        [10]   // MV 36,TEMPERATURE SETPOINT E. 1/10 DEGREE 'C'
        [12]   // MV 36,TEMPERATURE SETPOINT F. 1/10 DEGREE 'C'
        [14]   // MV 36,TEMPERATURE SETPOINT G. 1/10 DEGREE 'C'
        [13]   // MV 36,TEMPERATURE BREAKPOINT G. TIME 1/10 HOURS(ALWAYS=0)
        [15].2   // MV 36,PLC TO FOLLOW RAMP Breakpoints A to B
        [30].6   // MV 36,Current vessel cold cond.temp.reached
        [27]   // MV 36,CURRENT ELAPSED HOURS *10
        [30].5   // MV 36,Current vessel deferred chilling temp.high flag
        [1]   // MV 36,TEMPERATURE BREAKPOINT A. TIME 1/10 HOURS(ALWAYS=0)
        [29].1   // MV 36,Current vessel deferred chilling enabled flag
        [30].0   // MV 36,Cooling Valve to open
        [3]   // MV 36,TEMPERATURE BREAKPOINT B. TIME 1/10 HOURS(ALWAYS=0)
        [5]   // MV 36,TEMPERATURE BREAKPOINT C. TIME 1/10 HOURS(ALWAYS=0)
        [7]   // MV 36,TEMPERATURE BREAKPOINT D. TIME 1/10 HOURS(ALWAYS=0)
        [9]   // MV 36,TEMPERATURE BREAKPOINT E. TIME 1/10 HOURS(ALWAYS=0)
        [22]   // MV 36,Current FV total residence time
        [15].7   // MV 36,PC>PLC Rousing enabled
        [29].0   // MV 36,PC TO SAVE TEMPERATURE DATA
        [43]   // MV 36,Current vessel powder type
        [44]   // MV 36,Current vessel powder amount
        [15].3   // MV 36,PLC TO USE CONE COOLING JACKET
        [25]   // MV 36,ACTUAL TEMPERATURE -DEGREES 'C'*10
        [15]   // MV 36,FLAGS-PROFILE CONTROL
        [26]   // MV 36,Calculated Setpoint 1/10 degrees C
        [20]   // MV 36,Current FV warm conditioning time
        [29]   // MV 36,FLAGS - PLC CONTROL
        [30].1   // MV 36,Rouser required
        [28]   // MV 36,CURRENT VOLUME HL*10
   MV_N151 : INT[50] := ([0] := 347, [2] := 100, [3] := 1200, [4] := 100, [5] := 1680, [6] := -15, [7] := 5280, [8] := -15, [9] := 7210, [10] := -15, [11] := 8340, [12] := -15, [13] := 32767, [14] := -15, [15] := 164, [17] := -32767, [18] := -32767, [19] := 1680, [20] := 1200, [21] := 2981, [22] := 6282, [23] := 1, [24] := 13, [25] := -12, [26] := -15, [27] := 4630, [30] := 123, [32] := 2, [34] := 2, [40] := 2);   // MV 47, CURRENT FV DATA
        [24]   // MV 47,Phase 0=off 8=Wait yeast 9=Wait Fill 10=Maturation 11to16=Conditioning
        [15].9   // MV 47,Current vessel deferred chilling manual override
        [15].4   // MV 47,Profile Control Flags : This is a Maturation Profile
        [30].3   // MV 47,Current vessel deferred chilling active
        [15].5   // MV 47,Profile Control Flags : This is a Conditioning Profile
        [11]   // MV 47,TEMPERATURE BREAKPOINT F. TIME 1/10 HOURS(ALWAYS=0)
        [13]   // MV 47,TEMPERATURE BREAKPOINT G. TIME 1/10 HOURS(ALWAYS=0)
        [16].1   // MV 47,Profile control flag Hold at B.P B
        [16].2   // MV 47,Profile control flag Hold at B.P C
        [16].3   // MV 47,Profile control flag Hold at B.P D
        [30].5   // MV 47,Current vessel deferred chilling temp.high flag
        [36]   // MV 47,Current vessel time to deferred chlling start (hrs.x10)
        [16].4   // MV 47,Profile control flag Hold at B.P E
        [16].5   // MV 47,Profile control flag Hold at B.P F
        [16].6   // MV 47,Profile control flag Hold at B.P G
        [0]   // MV 47,FV SYSTEM WORKING BUFFER VESSEL NUMBER
        [21]   // MV 47,Current vessel cold conditioning time
        [2]   // MV 47,TEMPERATURE SETPOINT A. 1/10 DEGREE 'C'
        [30].4   // MV 47,Current vessel final temp.reached
        [4]   // MV 47,TEMPERATURE SETPOINT B. 1/10 DEGREE 'C'
        [6]   // MV 47,TEMPERATURE SETPOINT C. 1/10 DEGREE 'C'
        [8]   // MV 47,TEMPERATURE SETPOINT D. 1/10 DEGREE 'C'
        [40]   // MV 47,Vessel RoutingStatus 0=Clean,1=Filling,2= Beer,3=Packng1,4=Pac kng2,5=Packng3,6=Ven ting,7=Dirty,8=CIP
        [10]   // MV 47,TEMPERATURE SETPOINT E. 1/10 DEGREE 'C'
        [1]   // MV 47,TEMPERATURE BREAKPOINT A. TIME 1/10 HOURS(ALWAYS=0)
        [12]   // MV 47,TEMPERATURE SETPOINT F. 1/10 DEGREE 'C'
        [14]   // MV 47,TEMPERATURE SETPOINT G. 1/10 DEGREE 'C'
        [29].1   // MV 47,Current vessel deferred chilling enabled flag
        [15].2   // MV 47,PLC TO FOLLOW RAMP Breakpoints A to B
        [30].6   // MV 47,Current vessel cold cond.temp.reached
        [3]   // MV 47,TEMPERATURE BREAKPOINT B. TIME 1/10 HOURS(ALWAYS=0)
        [5]   // MV 47,TEMPERATURE BREAKPOINT C. TIME 1/10 HOURS(ALWAYS=0)
        [27]   // MV 47,CURRENT ELAPSED HOURS *10
        [30].0   // MV 47,Cooling Valve to open
        [7]   // MV 47,TEMPERATURE BREAKPOINT D. TIME 1/10 HOURS(ALWAYS=0)
        [9]   // MV 47,TEMPERATURE BREAKPOINT E. TIME 1/10 HOURS(ALWAYS=0)
        [22]   // MV 47,Current FV total residence time
        [15].7   // MV 47,PC>PLC Rousing enabled
        [43]   // MV 47,Current vessel powder type
        [29].0   // MV 47,PC TO SAVE TEMPERATURE DATA
        [15].3   // MV 47,PLC TO USE CONE COOLING JACKET
        [44]   // MV 47,Current vessel powder amount
        [25]   // MV 47,ACTUAL TEMPERATURE -DEGREES 'C'*10
        [15]   // MV 47,FLAGS-PROFILE CONTROL
        [26]   // MV 47,Calculated Setpoint 1/10 degrees C
        [20]   // MV 47,Current FV warm conditioning time
        [29]   // MV 47,FLAGS - PLC CONTROL
        [30].1   // MV 47,Rouser required
        [28]   // MV 47,CURRENT VOLUME HL*10
   MV_N15_63_0_OutputBit : BOOL;
   MV_N190 : INT[255] := ([0] := 1, [2] := 2, [3] := 2, [4] := 7, [5] := 2, [6] := 2, [7] := 2, [8] := 2, [9] := 2, [10] := 7, [11] := 7, [12] := 7, [13] := 2, [100] := 1, [101] := 2048, [102] := 10, [103] := 14, [105] := 13, [106] := 10, [107] := 15, [108] := 10, [109] := 10, [113] := 10, [200] := 8194, [201] := -16384, [203] := 20, [204] := 11, [205] := 137, [206] := 100, [209] := 23, [215] := 14641, [216] := 11826, [217] := 13873, [218] := 11832, [219] := 12338, [220] := 13102, [221] := 52);   // Original N File From SLC, No Description Available
        [200].0   // Heartbeat Fault
        [101].0   // MV36 Rouser On to Remote I/O on MV Routing PLC
        [101].1   // MV37 Rouser On to Remote I/O on MV Routing PLC
        [101].2   // MV38 Rouser On to Remote I/O on MV Routing PLC
        [101].3   // MV39 Rouser On to Remote I/O on MV Routing PLC
        [101].4   // MV40 Rouser On to Remote I/O on MV Routing PLC
        [101].5   // MV41 Rouser On to Remote I/O on MV Routing PLC
        [101].6   // MV42 Rouser On to Remote I/O on MV Routing PLC
        [101].7   // MV43 Rouser On to Remote I/O on MV Routing PLC
        [101].10   // MV46 Rouser On to Remote I/O on MV Routing PLC
        [101].11   // MV47 Rouser On to Remote I/O on MV Routing PLC
        [101].8   // MV44 Rouser On to Remote I/O on MV Routing PLC
        [101].9   // MV45 Rouser On to Remote I/O on MV Routing PLC
        [102]   // MV36 Ageing Status to Routing PLC
        [103]   // MV37 Ageing Status to Routing PLC
        [104]   // MV46 Ageing Status to Routing PLC
        [105]   // MV47 Ageing Status to Routing PLC
        [106]   // MV38 Ageing Status to Routing PLC
        [107]   // MV39 Ageing Status to Routing PLC
        [108]   // MV40 Ageing Status to Routing PLC
        [109]   // MV41 Ageing Status to Routing PLC
        [110]   // MV42 Ageing Status to Routing PLC
        [111]   // MV43 Ageing Status to Routing PLC
        [112]   // MV44 Ageing Status to Routing PLC
        [100].0   // MV Aging (This) PLC Heartbeat
        [1]   // Rouser Feedbacks from MV Routing PLC
        [113]   // MV45 Ageing Status to Routing PLC
        [200].1   // Enable Comms to MV Routing PLC
        [2]   // MV36 Routing Status from Routing PLC
        [3]   // MV37 Routing Status from Routing PLC
        [201]   // Comms to MV Routing PLC
        [4]   // MV46 Routing Status from Routing PLC
        [5]   // MV47 Routing Status from Routing PLC
        [0].0   // MV Routing PLC Heartbeat
   MV_N255 : DINT[255] := ([0] := 1536, [1] := 2048, [2] := 2048, [3] := 2048, [4] := 2048, [5] := 2048, [6] := 2048, [7] := 1536, [8] := 2048, [9] := 2048, [10] := 2048, [11] := 1536, [12] := 2048, [13] := 2048, [14] := 2048, [15] := 2048, [16] := 1536, [17] := 2048, [18] := 2048, [19] := 2048, [20] := 2048, [21] := 2048, [22] := 2048, [23] := 2048, [24] := 2048, [25] := 1536, [26] := 2048, [27] := 1536, [28] := 2048, [32] := 17984, [33] := 2112, [34] := 2112, [35] := 2112, [36] := 2112, [37] := 2112, [38] := 2112, [39] := 2112, [40] := 2112, [41] := 2112, [42] := 2112, [43] := 2112, [44] := 2112, [45] := 2112, [46] := 2112, [47] := 2112, [48] := 2112, [49] := 2112, [50] := 2112, [51] := 2112, [52] := 2112, [53] := 2112, [54] := 2112, [55] := 2112, [56] := 2112, [57] := 2368, [58] := 2112, [59] := 2368, [60] := 2112, [64] := 2048, [65] := 2048,
        [66] := 2048, [67] := 2048, [68] := 2048, [69] := 2048, [70] := 2048, [71] := 2048, [72] := 2048, [73] := 2048, [74] := 2048, [75] := 1536);   // Old Format Checkwords To Keep Delphi Indicating Status Correctly.
   MV_N7 : INT[255] := ([0] := 2);   // INTEGER
        [0]   // Temp.register
   MV_Old_CW_Num : DINT;
   MV_SFile : INT[255] := ([37] := 2020, [40] := 17, [42] := 5);   // SLC Equivalent System File, So Original Code Can Remain
        [41]   // Clock Calendar Minutes
        [42]   // Clock Calendar Seconds
        [1].15   // First Scan Flag
        [13]   // Remainder Result From Divide
        [37]   // Clock System Year
        [40]   // Clock Calendar Hours
   MV_T102 : TIMER[10] := ([0].PRE := 360000, [0].ACC := 260086, [0].EN := 1, [0].TT := 1);
   MV_T16 : TIMER[10] := ([0].PRE := 3000, [0].ACC := 330, [0].EN := 1, [0].TT := 1);
   MV_T191 : TIMER[20] := ([0].PRE := 20000, [1].PRE := 20000, [1].ACC := 741, [1].EN := 1, [1].TT := 1);
   MV_T4 : TIMER[20] := ([2].PRE := 1000, [2].ACC := 177, [2].EN := 1, [2].TT := 1);
   MV_TENTH_HOUR_OUTPUT_BIT : BOOL;
   MV_to_data_file : DINT;
   MV_to_data_offset : DINT;
   MV_TP_CaskEmptyingPressure : REAL := 3.0;
   MV_TP_CaskFillingPressure : REAL := 3.0;
   MV_TP_CaskPrefillPressure : REAL := 1.0;
   MV_TP_CaskStoragePressure : REAL := 4.0;
   MV_TP_CaskStoragePressureDelay : DINT := 48;
   MV_TP_CaskStoragePressureDelay_Secs : DINT := 43200;
   MV_TP_CaskStoragePressureLevel : REAL := 170.0;
   MV_TP_DALChase_Time : DINT := 90000;
   MV_TP_Deadband : REAL := 1.0;
   MV_TP_Emptying_Volume_Setpoint : REAL := 250.0;
   MV_TP_HighLevelDeadband : REAL := 2.0;
   MV_TP_HighLevelDeadband_1 : REAL := 2.0;
   MV_TP_KBEmptyingPressure : REAL := 15.0;
   MV_TP_KBFillingPressure : REAL := 3.0;
   MV_TP_KBPrefillPressure : REAL := 2.5;
   MV_TP_KBPurgeTime : DINT;
   MV_TP_KBStoragePressure : REAL := 10.0;
   MV_TP_KBStoragePressureLevel : REAL := 200.0;
   MV_TP_LowLevelDeadbandThreshold : REAL;
   MV_TP_LowLevelDeadbandThreshold_1 : REAL := 0.3;
   MV_TP_NoCIPDelay : DINT;
   MV_TP_OtherVesselsNotVentingDelay : DINT;
   MV_TP_VentPressure : REAL := 0.3;
   MV_value_to_set : INT;
   MV_WarningTimeout : DINT;
   MV_word_offset : INT := 24;
   MVCT_Proxies_OK : BOOL;
   MVCT_ProxiesCIP_OK : DINT;
   New_Item : PlantItem := (CW := 2#0000_0000_0000_0000_0010_0010_0100_0001, DriveBits := 1);
   new_item_temp : DINT := 385;
   Old_Item : INT := 385;
   old_item_bit_mask : DINT := 19968;
   old_item_temp : DINT := 8769;
   One_Minute_One_Scan : BOOL;
   One_Minute_One_Scan_Timer : TIMER := (PRE := 60000, ACC := 22669, EN := 1, TT := 1);
   One_sec_toggle : DINT;
   One_Second_1_scan : BOOL;
   One_Second_One_Scan : ALIAS FOR One_Second_1_scan;
   One_Second_Toggle : BOOL := 1;
   One_Second_Toggle_Valid_Groups : BOOL := 1;
   overrange_RIO_analog_value : REAL;
   pe_test : DINT := 55;
   pe_test2 : DINT := 2;
   rack_simulation_flag : BOOL := 1;
   reset_msg_interval : BOOL;
   result_string : STRING := '989:42:05';
   Scada_Pump_Fault_No : DINT := 20001;
   Scada_Pump_H_Fault_No : DINT := 20001;
   Scada_Pump_T_Fault_No : DINT := 20001;
   Scada_Valve_Fault_No : DINT;
   scada_watchdog : DINT := 29;
   scale_analog_int : DINT;
   scale_analog_result : REAL := 150.0;
   scale_eu_max : REAL := 20000.0;
   scale_eu_min : REAL;
   scale_raw_input : REAL;
   scale_raw_max : REAL := 100.0;
   scale_raw_min : REAL;
   scale_routine_active : BOOL := 1;
   scale_temp : REAL := 160.0;
   se_string : STRING := '6';
   seconds_input : INT;
   seconds_input_DINT : DINT := 3562924;
   temp : INT := 984;
   temp_counter : DINT := 23;
   temp_hr : INT;
   temp_mn : INT := 42;
   temp_se : INT := 4;
   TempChecktime : DINT := 64;
   template_analog_input : PlantItem;
   template_analog_input_RawInput : REAL;
   template_analog_output : PlantItem;
   template_analog_output_RawOutput : REAL;
   template_boolean : BOOL;
   template_input : PlantItem;
   template_input_RawInput : ALIAS FOR template_boolean;
   template_output : PlantItem;
   template_output_RawOutput : ALIAS FOR template_boolean;   // P04CHILLRUN Chiller Run Signal
   template_pump : PlantItem;
   template_pump_D : ALIAS FOR template_boolean;   // auto start vacuum pump 1
   template_pump_H : ALIAS FOR template_boolean;   // vacuum pump 1 auto avail
   template_pump_ISOL : ALIAS FOR template_boolean;
   template_pump_R : ALIAS FOR template_boolean;   // vacuum pump 1 running
   template_valve : PlantItem;
   template_valve_C : ALIAS FOR template_boolean;   // skim manifold to ycv2 drain valve closed
   template_valve_DR : ALIAS FOR template_boolean;   // drive open skim manifold to ycv2 drain valve
   template_valve_O : ALIAS FOR template_boolean;   // skim manifold to ycv2 drain valve opened
   test : INT := -32767;
   test_alm : BOOL;
   test_alm_out : BOOL;
   testing_bit : BOOL := 1;
   underrange_RIO_analog_value : REAL;
   Unused_Healthy_Feedback : BOOL := 1;
   Unused_NotTripped_Feedback : BOOL := 1;
   YST_Data : REAL[2] := ([0] := 134.1, [1] := 140.96251);
   zero_string : STRING := '0'; {constant, access Read Only}
END_VAR

PROGRAM _1Second   (* main routine OneSecond *)

ROUTINE OneSecond   (* ladder *)
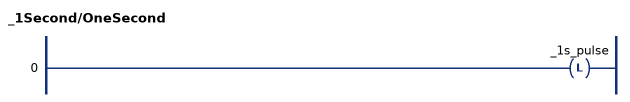
   0: OTL(_1s_pulse);
END_ROUTINE
END_PROGRAM

PROGRAM First_Task   (* main routine MainRoutine *)

ROUTINE MainRoutine   (* ladder *)
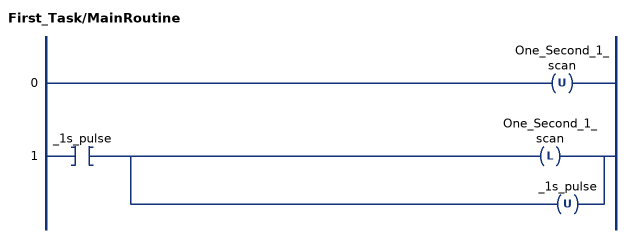
   0: OTU(One_Second_1_scan);
   1: XIC(_1s_pulse)[OTL(One_Second_1_scan) ,OTU(_1s_pulse) ];
END_ROUTINE
END_PROGRAM

PROGRAM Last_Task   (* main routine MainRoutine *)

ROUTINE MainRoutine   (* ladder *)
   0: NOP();
END_ROUTINE
END_PROGRAM

PROGRAM MC_Common   (* main routine MC_MAIN *)
VAR
   MC_CH2_CIP_BYPASS_CIP : BOOL := 1;
   MC_CIP_String_Result1 : DINT;
   MC_CIP_String_Result2 : DINT;
   MC_CIP_String_Result3 : DINT;
   MC_CIP_String_Result4 : DINT;
   MC_CIP_String_Result5 : DINT;
   MC_CIP_String_Result6 : DINT;
END_VAR

ROUTINE A_FactoryTalk_Requirements   (* ladder *)
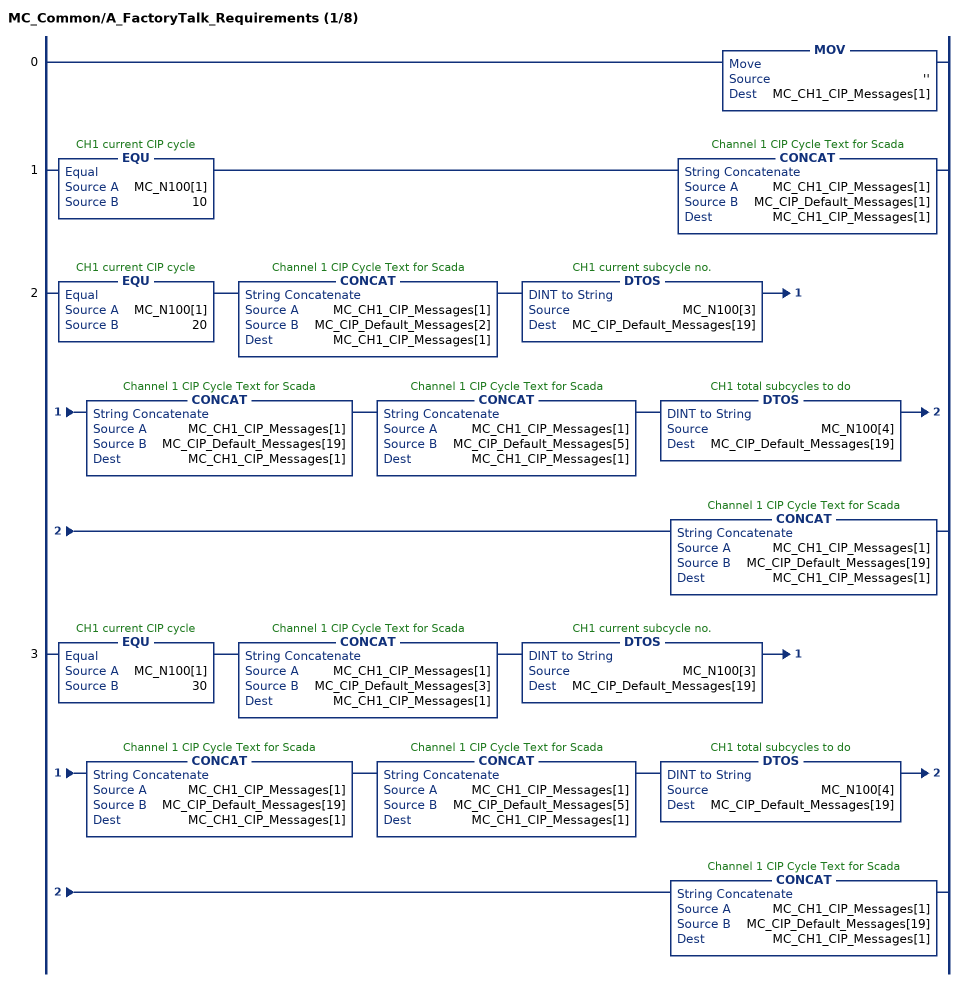
   0: MOV('',MC_CH1_CIP_Messages[1]);
   1: EQU(MC_N100[1],10)CONCAT(MC_CH1_CIP_Messages[1],MC_CIP_Default_Messages[1],MC_CH1_CIP_Messages[1]);
   2: EQU(MC_N100[1],20)CONCAT(MC_CH1_CIP_Messages[1],MC_CIP_Default_Messages[2],MC_CH1_CIP_Messages[1])DTOS(MC_N100[3],MC_CIP_Default_Messages[19])CONCAT(MC_CH1_CIP_Messages[1],MC_CIP_Default_Messages[19],MC_CH1_CIP_Messages[1])CONCAT(MC_CH1_CIP_Messages[1],MC_CIP_Default_Messages[5],MC_CH1_CIP_Messages[1])DTOS(MC_N100[4],MC_CIP_Default_Messages[19])CONCAT(MC_CH1_CIP_Messages[1],MC_CIP_Default_Messages[19],MC_CH1_CIP_Messages[1]);
   3: EQU(MC_N100[1],30)CONCAT(MC_CH1_CIP_Messages[1],MC_CIP_Default_Messages[3],MC_CH1_CIP_Messages[1])DTOS(MC_N100[3],MC_CIP_Default_Messages[19])CONCAT(MC_CH1_CIP_Messages[1],MC_CIP_Default_Messages[19],MC_CH1_CIP_Messages[1])CONCAT(MC_CH1_CIP_Messages[1],MC_CIP_Default_Messages[5],MC_CH1_CIP_Messages[1])DTOS(MC_N100[4],MC_CIP_Default_Messages[19])CONCAT(MC_CH1_CIP_Messages[1],MC_CIP_Default_Messages[19],MC_CH1_CIP_Messages[1]);
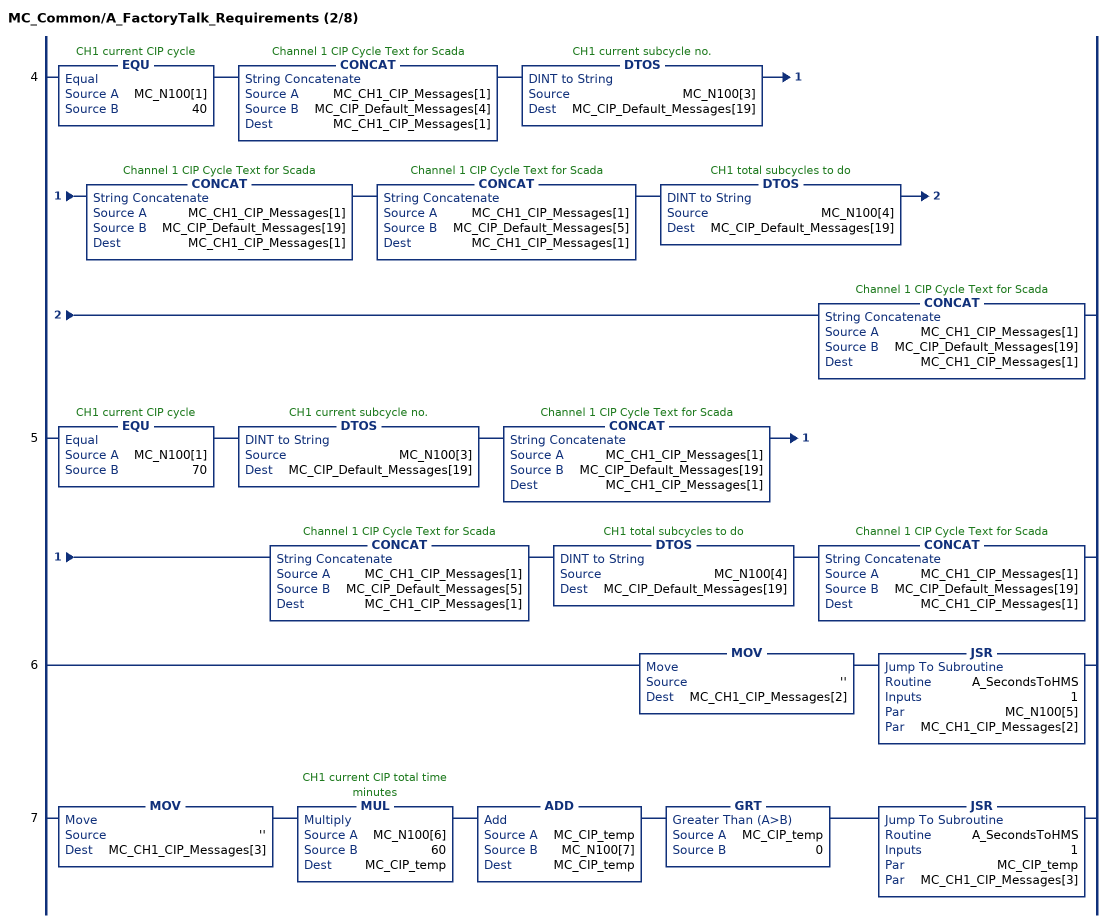
   4: EQU(MC_N100[1],40)CONCAT(MC_CH1_CIP_Messages[1],MC_CIP_Default_Messages[4],MC_CH1_CIP_Messages[1])DTOS(MC_N100[3],MC_CIP_Default_Messages[19])CONCAT(MC_CH1_CIP_Messages[1],MC_CIP_Default_Messages[19],MC_CH1_CIP_Messages[1])CONCAT(MC_CH1_CIP_Messages[1],MC_CIP_Default_Messages[5],MC_CH1_CIP_Messages[1])DTOS(MC_N100[4],MC_CIP_Default_Messages[19])CONCAT(MC_CH1_CIP_Messages[1],MC_CIP_Default_Messages[19],MC_CH1_CIP_Messages[1]);
   5: EQU(MC_N100[1],70)DTOS(MC_N100[3],MC_CIP_Default_Messages[19])CONCAT(MC_CH1_CIP_Messages[1],MC_CIP_Default_Messages[19],MC_CH1_CIP_Messages[1])CONCAT(MC_CH1_CIP_Messages[1],MC_CIP_Default_Messages[5],MC_CH1_CIP_Messages[1])DTOS(MC_N100[4],MC_CIP_Default_Messages[19])CONCAT(MC_CH1_CIP_Messages[1],MC_CIP_Default_Messages[19],MC_CH1_CIP_Messages[1]);
   6: MOV('',MC_CH1_CIP_Messages[2])JSR(A_SecondsToHMS,1,MC_N100[5],MC_CH1_CIP_Messages[2]);
   7: MOV('',MC_CH1_CIP_Messages[3])MUL(MC_N100[6],60,MC_CIP_temp)ADD(MC_CIP_temp,MC_N100[7],MC_CIP_temp)GRT(MC_CIP_temp,0)JSR(A_SecondsToHMS,1,MC_CIP_temp,MC_CH1_CIP_Messages[3]);
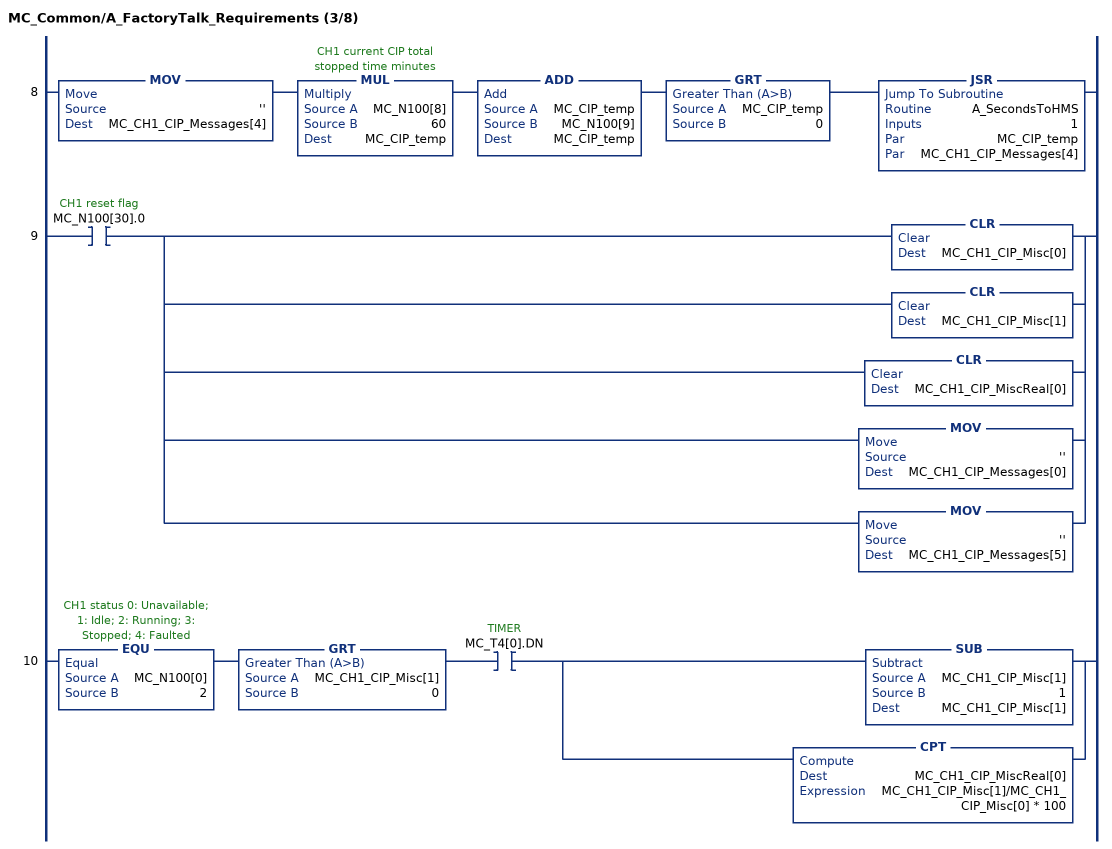
   8: MOV('',MC_CH1_CIP_Messages[4])MUL(MC_N100[8],60,MC_CIP_temp)ADD(MC_CIP_temp,MC_N100[9],MC_CIP_temp)GRT(MC_CIP_temp,0)JSR(A_SecondsToHMS,1,MC_CIP_temp,MC_CH1_CIP_Messages[4]);
   9: XIC(MC_N100[30].0)[CLR(MC_CH1_CIP_Misc[0]) ,CLR(MC_CH1_CIP_Misc[1]) ,CLR(MC_CH1_CIP_MiscReal[0]) ,MOV('',MC_CH1_CIP_Messages[0]) ,MOV('',MC_CH1_CIP_Messages[5]) ];
   10: EQU(MC_N100[0],2)GRT(MC_CH1_CIP_Misc[1],0)XIC(MC_T4[0].DN)[SUB(MC_CH1_CIP_Misc[1],1,MC_CH1_CIP_Misc[1]) ,CPT(MC_CH1_CIP_MiscReal[0],MC_CH1_CIP_Misc[1]/MC_CH1_CIP_Misc[0] * 100) ];
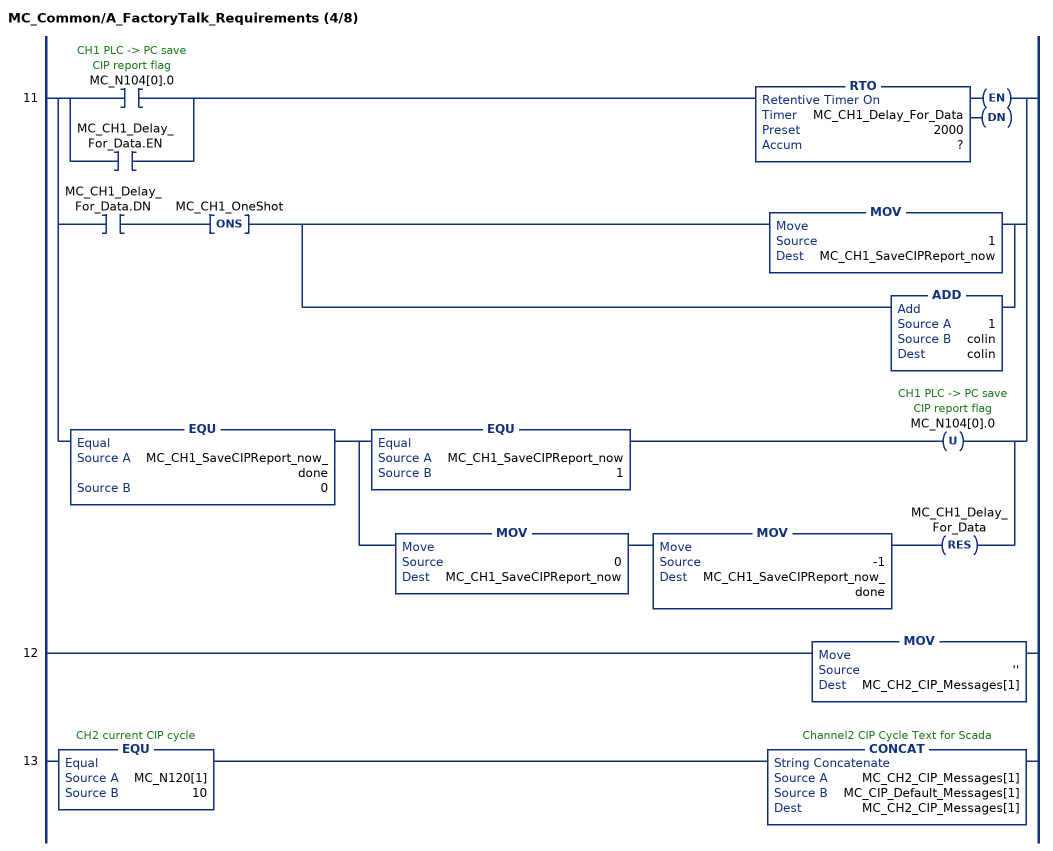
   11: [[XIC(MC_N104[0].0) ,XIC(MC_CH1_Delay_For_Data.EN) ] RTO(MC_CH1_Delay_For_Data,?,?) ,XIC(MC_CH1_Delay_For_Data.DN) ONS(MC_CH1_OneShot) [MOV(1,MC_CH1_SaveCIPReport_now) ,ADD(1,colin,colin) ] ,EQU(MC_CH1_SaveCIPReport_now_done,0) [EQU(MC_CH1_SaveCIPReport_now,1) OTU(MC_N104[0].0) ,MOV(0,MC_CH1_SaveCIPReport_now) MOV(-1,MC_CH1_SaveCIPReport_now_done) RES(MC_CH1_Delay_For_Data) ] ];
   12: MOV('',MC_CH2_CIP_Messages[1]);
   13: EQU(MC_N120[1],10)CONCAT(MC_CH2_CIP_Messages[1],MC_CIP_Default_Messages[1],MC_CH2_CIP_Messages[1]);
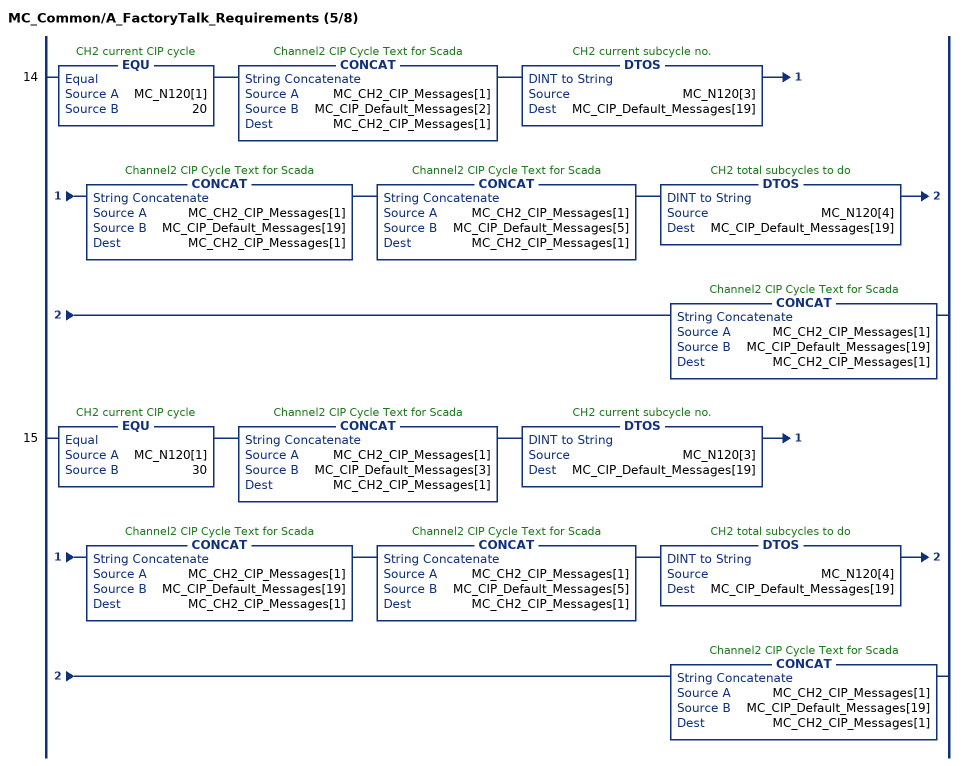
   14: EQU(MC_N120[1],20)CONCAT(MC_CH2_CIP_Messages[1],MC_CIP_Default_Messages[2],MC_CH2_CIP_Messages[1])DTOS(MC_N120[3],MC_CIP_Default_Messages[19])CONCAT(MC_CH2_CIP_Messages[1],MC_CIP_Default_Messages[19],MC_CH2_CIP_Messages[1])CONCAT(MC_CH2_CIP_Messages[1],MC_CIP_Default_Messages[5],MC_CH2_CIP_Messages[1])DTOS(MC_N120[4],MC_CIP_Default_Messages[19])CONCAT(MC_CH2_CIP_Messages[1],MC_CIP_Default_Messages[19],MC_CH2_CIP_Messages[1]);
   15: EQU(MC_N120[1],30)CONCAT(MC_CH2_CIP_Messages[1],MC_CIP_Default_Messages[3],MC_CH2_CIP_Messages[1])DTOS(MC_N120[3],MC_CIP_Default_Messages[19])CONCAT(MC_CH2_CIP_Messages[1],MC_CIP_Default_Messages[19],MC_CH2_CIP_Messages[1])CONCAT(MC_CH2_CIP_Messages[1],MC_CIP_Default_Messages[5],MC_CH2_CIP_Messages[1])DTOS(MC_N120[4],MC_CIP_Default_Messages[19])CONCAT(MC_CH2_CIP_Messages[1],MC_CIP_Default_Messages[19],MC_CH2_CIP_Messages[1]);
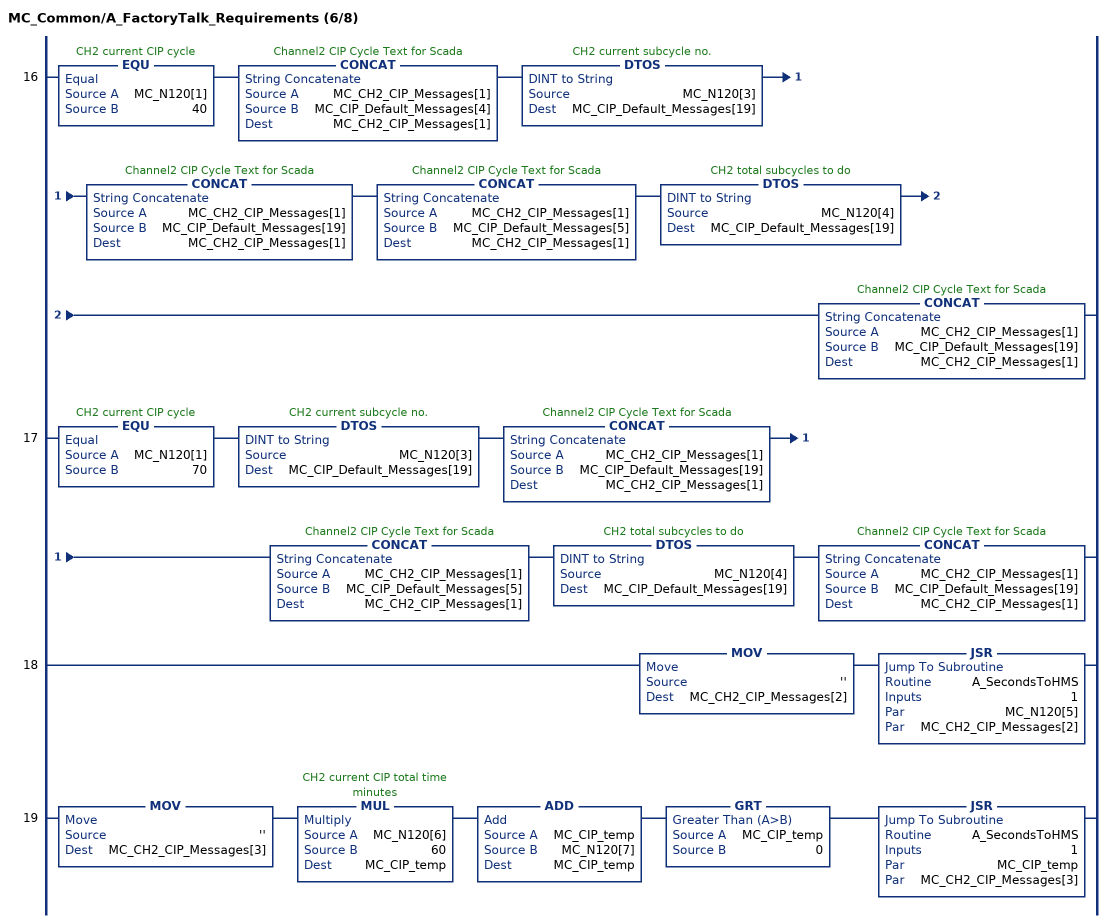
   16: EQU(MC_N120[1],40)CONCAT(MC_CH2_CIP_Messages[1],MC_CIP_Default_Messages[4],MC_CH2_CIP_Messages[1])DTOS(MC_N120[3],MC_CIP_Default_Messages[19])CONCAT(MC_CH2_CIP_Messages[1],MC_CIP_Default_Messages[19],MC_CH2_CIP_Messages[1])CONCAT(MC_CH2_CIP_Messages[1],MC_CIP_Default_Messages[5],MC_CH2_CIP_Messages[1])DTOS(MC_N120[4],MC_CIP_Default_Messages[19])CONCAT(MC_CH2_CIP_Messages[1],MC_CIP_Default_Messages[19],MC_CH2_CIP_Messages[1]);
   17: EQU(MC_N120[1],70)DTOS(MC_N120[3],MC_CIP_Default_Messages[19])CONCAT(MC_CH2_CIP_Messages[1],MC_CIP_Default_Messages[19],MC_CH2_CIP_Messages[1])CONCAT(MC_CH2_CIP_Messages[1],MC_CIP_Default_Messages[5],MC_CH2_CIP_Messages[1])DTOS(MC_N120[4],MC_CIP_Default_Messages[19])CONCAT(MC_CH2_CIP_Messages[1],MC_CIP_Default_Messages[19],MC_CH2_CIP_Messages[1]);
   18: MOV('',MC_CH2_CIP_Messages[2])JSR(A_SecondsToHMS,1,MC_N120[5],MC_CH2_CIP_Messages[2]);
   19: MOV('',MC_CH2_CIP_Messages[3])MUL(MC_N120[6],60,MC_CIP_temp)ADD(MC_CIP_temp,MC_N120[7],MC_CIP_temp)GRT(MC_CIP_temp,0)JSR(A_SecondsToHMS,1,MC_CIP_temp,MC_CH2_CIP_Messages[3]);
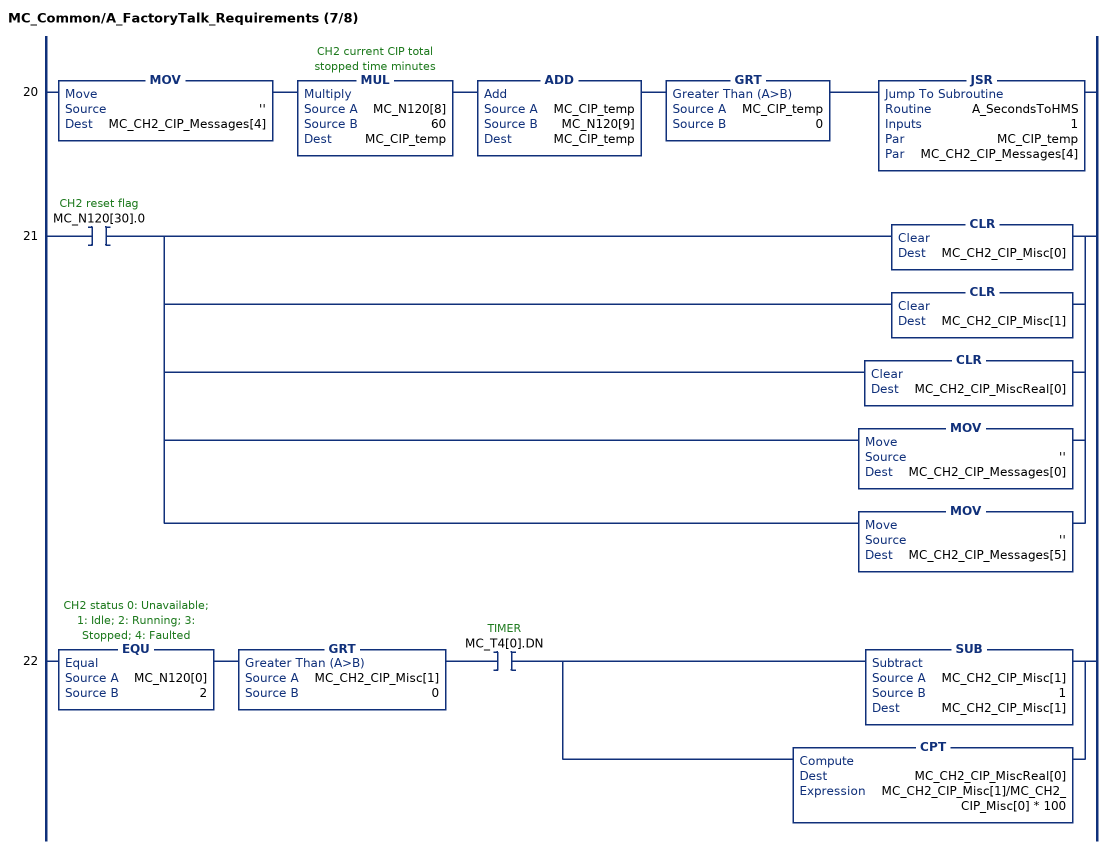
   20: MOV('',MC_CH2_CIP_Messages[4])MUL(MC_N120[8],60,MC_CIP_temp)ADD(MC_CIP_temp,MC_N120[9],MC_CIP_temp)GRT(MC_CIP_temp,0)JSR(A_SecondsToHMS,1,MC_CIP_temp,MC_CH2_CIP_Messages[4]);
   21: XIC(MC_N120[30].0)[CLR(MC_CH2_CIP_Misc[0]) ,CLR(MC_CH2_CIP_Misc[1]) ,CLR(MC_CH2_CIP_MiscReal[0]) ,MOV('',MC_CH2_CIP_Messages[0]) ,MOV('',MC_CH2_CIP_Messages[5]) ];
   22: EQU(MC_N120[0],2)GRT(MC_CH2_CIP_Misc[1],0)XIC(MC_T4[0].DN)[SUB(MC_CH2_CIP_Misc[1],1,MC_CH2_CIP_Misc[1]) ,CPT(MC_CH2_CIP_MiscReal[0],MC_CH2_CIP_Misc[1]/MC_CH2_CIP_Misc[0] * 100) ];
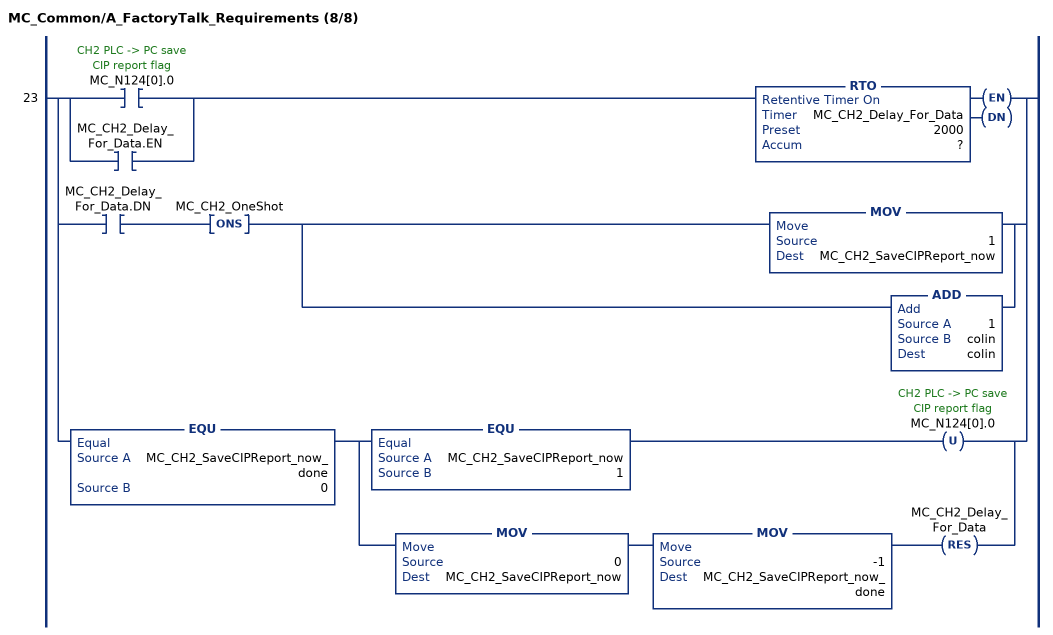
   23: [[XIC(MC_N124[0].0) ,XIC(MC_CH2_Delay_For_Data.EN) ] RTO(MC_CH2_Delay_For_Data,?,?) ,XIC(MC_CH2_Delay_For_Data.DN) ONS(MC_CH2_OneShot) [MOV(1,MC_CH2_SaveCIPReport_now) ,ADD(1,colin,colin) ] ,EQU(MC_CH2_SaveCIPReport_now_done,0) [EQU(MC_CH2_SaveCIPReport_now,1) OTU(MC_N124[0].0) ,MOV(0,MC_CH2_SaveCIPReport_now) MOV(-1,MC_CH2_SaveCIPReport_now_done) RES(MC_CH2_Delay_For_Data) ] ];
END_ROUTINE

ROUTINE A_SecondsToHMS   (* ladder *)
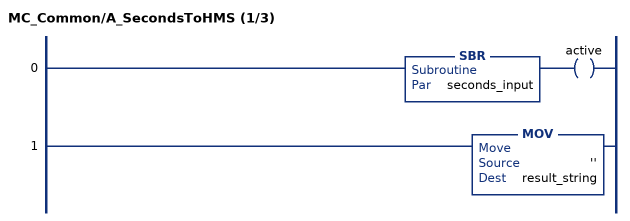
   0: SBR(seconds_input)OTE(active);
   1: MOV('',result_string);
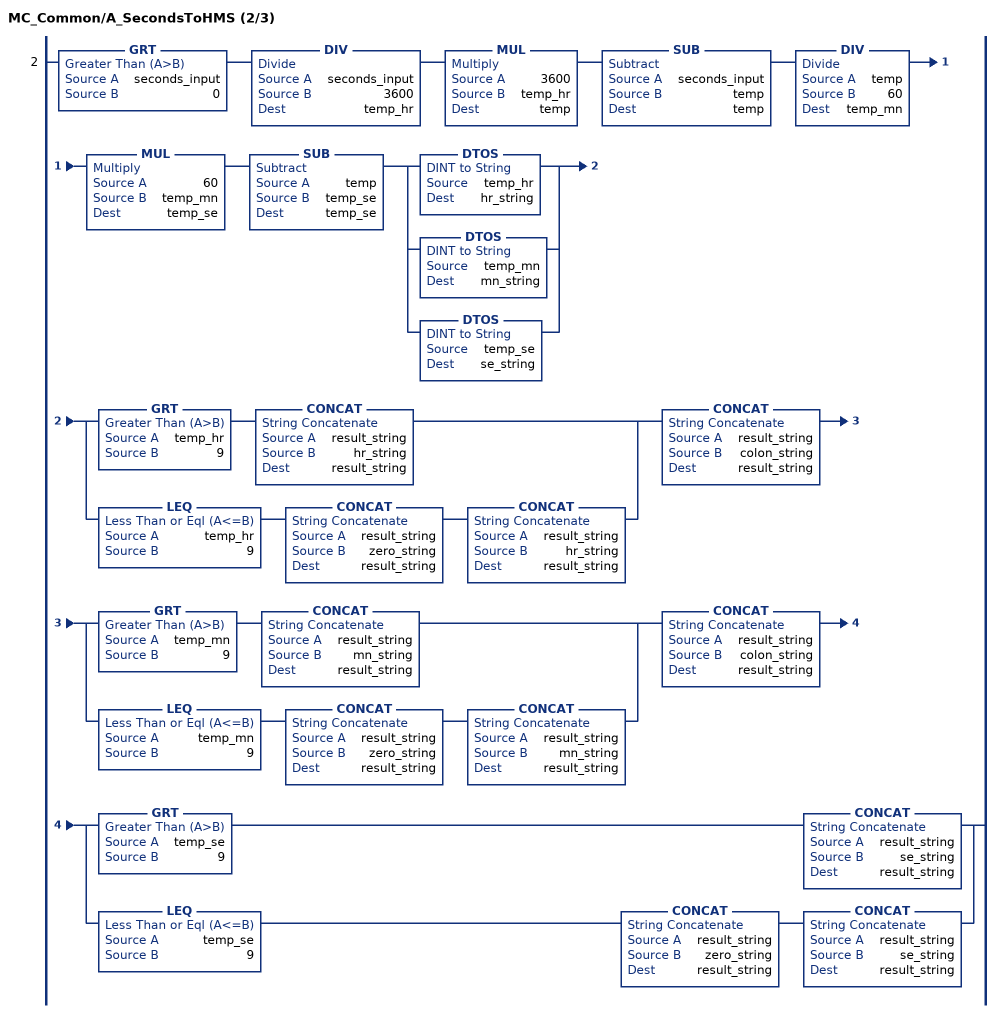
   2: GRT(seconds_input,0)DIV(seconds_input,3600,temp_hr)MUL(3600,temp_hr,temp)SUB(seconds_input,temp,temp)DIV(temp,60,temp_mn)MUL(60,temp_mn,temp_se)SUB(temp,temp_se,temp_se)[DTOS(temp_hr,hr_string) ,DTOS(temp_mn,mn_string) ,DTOS(temp_se,se_string) ][GRT(temp_hr,9) CONCAT(result_string,hr_string,result_string) ,LEQ(temp_hr,9) CONCAT(result_string,zero_string,result_string) CONCAT(result_string,hr_string,result_string) ]CONCAT(result_string,colon_string,result_string)[GRT(temp_mn,9) CONCAT(result_string,mn_string,result_string) ,LEQ(temp_mn,9) CONCAT(result_string,zero_string,result_string) CONCAT(result_string,mn_string,result_string) ]CONCAT(result_string,colon_string,result_string)[GRT(temp_se,9) CONCAT(result_string,se_string,result_string) ,LEQ(temp_se,9) CONCAT(result_string,zero_string,result_string) CONCAT(result_string,se_string,result_string) ];
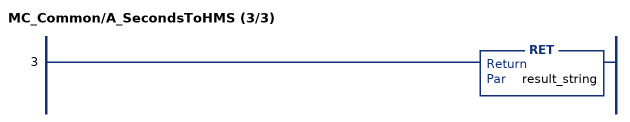
   3: RET(result_string);
END_ROUTINE
